      ProcessValue <- "Sequence Times_DB_Dwell Timer_Hours Left"
   IOField "I/O field_66" at 316,321 size 33x28; Authorization "User administration"; FormatPattern 99; Unit d
      ProcessValue <- "Sequence Times_DB_Dwell Timer_Days Left"
   IOField "I/O field_2" at 216,355 size 79x28; Authorization "Commissioning"; FormatPattern 999.9; Unit  Hrs
      ProcessValue <- "Sequence Times_DB_Re-Ox Time"
   IOField "I/O field_67" at 380,355 size 35x28; Authorization "User administration"; FormatPattern 99; Unit m
      ProcessValue <- "Sequence Times_DB_Re-Ox Timer_Minutes Left"
   IOField "I/O field_68" at 348,355 size 33x28; Authorization "User administration"; FormatPattern 99; Unit h
      ProcessValue <- "Sequence Times_DB_Re-Ox Timer_Hours Left"
   IOField "I/O field_69" at 316,355 size 33x28; Authorization "User administration"; FormatPattern 99; Unit d
      ProcessValue <- "Sequence Times_DB_Re-Ox Timer_Days Left"
   IOField "I/O field_70" at 216,389 size 79x28; Authorization "Commissioning"; FormatPattern 999.9; Unit  Hrs
      ProcessValue <- "Sequence Times_DB_Post-Dwell Time"
   IOField "I/O field_71" at 380,389 size 35x28; Authorization "User administration"; FormatPattern 99; Unit m
      ProcessValue <- "Sequence Times_DB_Post-Dwell Timer_Minutes Left"
   IOField "I/O field_72" at 348,389 size 33x28; Authorization "User administration"; FormatPattern 99; Unit h
      ProcessValue <- "Sequence Times_DB_Post-Dwell Timer_Hours Left"
   IOField "I/O field_73" at 316,389 size 33x28; Authorization "User administration"; FormatPattern 99; Unit d
      ProcessValue <- "Sequence Times_DB_Post-Dwell Timer_Days Left"
   Button "Button_1" at 364,1 size 56x38; TextOff 'Text'; PictureOff "Graphic_286"
      on Click: function_efd93a16("Tank Times", 300, 200, -1, -1, 1)
   Group "Group_1" at 20,501 size 235x37

PopupScreen "TANK Activ Warning" 665x250
   Button "Button_1" at 0,0 size 665x250; TextOff 'No TANK Selected. Select a TANK for Tank Treatment.'
      on Release: function_efd93a16("TANK Activ Warning", 300, 200, -1, -1, 1)
   Button "Button_2" at 208,187 size 250x35; TextOff 'OK, Select TANK'
      on Release: ActivateScreen("Balast Water Treatment Setup", 0); function_efd93a16("TANK Activ Warning", 0, 0, -1, -1, 1)

screen "Balast Water Treatment Plant Tank Pressure" 1280x800, template "Template"
   on GenerateScreen: "User_Change"(); "TitleUpdater"()
   Button "HmiScreenItemData_1" at 1,1 size 150x40; TextOn 'Back'; TextOff 'Main Index'
      on Release: ActivateScreen("02 Main Index", 0)
   TextField "Text field_63" at 383,107 size 72x30; Text 'Pre Dwell Time'
   Circle "Circle_29" at 1047,85 size 20x20
      Appearance <- "2102_TIME_CALCS_DB_POST_DWELL_TMR_DN"
   Button "HmiScreenItemData_9" at 10,60 size 158x27; TextOn 'Back'; TextOff 'BWTS Control'
   Button "HmiScreenItemData_4" at 14,150 size 75x47; TextOn 'Back'; TextOff 'Stop'; Authorization "Operate"
      on Release: function_efd93a16("BWTS Stop Confirm", 400, 200, -1, -1, 1)
      ObjectEnable <- "82_To_HMI_CRNT_MODE_GCU"
   Circle "Circle_20" at 137,105 size 29x29
      Appearance <- "80_From_HMI_RUN_IGG(1)"
   Button "HmiScreenItemData_3" at 14,93 size 75x47; TextOn 'Back'; TextOff 'Start'; Authorization "Operate"
      on Release: function_efd93a16("BWTS Start Confirm", 400, 200, -1, -1, 1)
      ObjectEnable <- "82_To_HMI_CRNT_MODE_GCU"
   Button "HmiScreenItemData_2" at 1129,1 size 150x40; TextOn 'Back'; TextOff 'BWTS Setup'
      on Release: ActivateScreen("Balast Water Treatment Setup", 0)
   TextField "Text field_1" at 290,107 size 68x30; Text 'Tank Selected'
   TextField "Text field_2" at 841,107 size 61x30; Text 'BWTS Started'
   TextField "Text field_3" at 568,107 size 62x30; Text 'IGGS Started'
   TextField "Text field_4" at 659,107 size 60x30; Text 'GCU Started'
   TextField "Text field_5" at 748,107 size 61x30; Text 'PGC Started'
   TextField "Text field_6" at 908,107 size 102x30; Text 'Gas Transfer Started'
   Circle "Circle_10" at 956,89 size 14x14
      Appearance <- "2110_BTCS_CNTRL_DB_BTCS_STEP"
   TextField "Text field_7" at 995,107 size 125x30; Text 'Treatment Cycle Completed'
   TextField "Text field_23" at 261,291 size 34x14; Text 'MBG'
   GraphicView "Graphic view_17" at 575,446 size 532x12; Picture "Graphic_151"
   Button "Button_13" at 252,437 size 37x30; TextOff 'DB&B'
   TextField "Text field_58" at 188,226 size 50x40; Text 'Safe Area'
   Button "Button_20" at 724,152 size 115x34; TextOff 'Re-Oxygenation'
      Appearance <- "2110_BTCS_CNTRL_DB_BTCS_STEP"
   Button "Button_21" at 845,152 size 93x34; TextOff 'Post Dwell'
      Appearance <- "2110_BTCS_CNTRL_DB_BTCS_STATE"
   Circle "Circle_1" at 137,105 size 29x29
      Appearance <- "2110_BTCS_CNTRL_DB_BTCS_STATE"
   Circle "Circle_8" at 775,89 size 14x14
      Appearance <- "2110_BTCS_CNTRL_DB_BTCS_STEP"
   Circle "Circle_9" at 685,89 size 14x14
      Appearance <- "100_GCU_AUTO_SEQ_DB_CRNT_STEP"
   Circle "Circle_11" at 595,89 size 14x14
      Appearance <- "51_SLAVE_STATUS_RUNNING"
   Circle "Circle_12" at 866,89 size 14x14
      Appearance <- "2110_BTCS_CNTRL_DB_BTCS_STEP"
   Circle "Circle_13" at 324,89 size 14x14
      Appearance <- "HMI Indication Logic_DB_Tank Selected"
   Circle "Circle_14" at 414,89 size 14x14
      Appearance <- "2102_TIME_CALCS_DB_PRE_DWELL_TMR_DN"
   Button "Button_3" at 626,152 size 93x34; TextOff 'Dwell'
      Appearance <- "2110_BTCS_CNTRL_DB_BTCS_STATE"
   Button "Button_5" at 944,152 size 93x34; TextOff 'Complete'
      Appearance <- "HMI Indication Logic_DB_Sequence Finished"
   TextField "Text field_61" at 202,107 size 71x30; Text 'FA Mode Selected'
   Circle "Circle_2" at 230,89 size 14x14
      Appearance <- "HMI Indication Logic_DB_FA Mode Selected"
   TextField "Text field_60" at 190,519 size 46x25; Text 'GCU'
   GraphicIOField "Graphic I/O field_4" at 187,543 size 53x55; PictureList "GCU"
      ProcessValue <- "100_GCU_AUTO_SEQ_DB_RNG"
   TextField "Text field_74" at 186,279 size 54x25; Text 'IGGS'
   GraphicIOField "Graphic I/O field_1" at 185,303 size 57x53; PictureList "IGGS"
      ProcessValue <- "14_DQ_Data_24PF1"
   TextField "Text field_62" at 183,359 size 60x20; Text 'Disabled'
   TextField "Text field_77" at 183,359 size 60x20; Text 'Enabled'
      Visibility <- "51_SLAVE_STATUS_RUNNING"
   Button "Button_8" at 178,280 size 70x105; TextOff 'Text'
      on Release: ActivateScreen("Inert Gas Generator Plant", 0)
   TextField "Text field_70" at 183,599 size 60x20; Text 'Disabled'
   TextField "Text field_71" at 183,599 size 60x20; Text 'Enabled'
      Visibility <- "100_GCU_AUTO_SEQ_DB_RNG"
   Button "Button_4" at 178,521 size 70x105; TextOff 'Text'
      on Release: ActivateScreen("Inert Gas Conditioning Plant", 0)
   GraphicIOField "Graphic I/O field_2" at 770,45 size 250x30; PictureList "Process time Banner"
      ProcessValue <- "2110_BTCS_CNTRL_DB_BTCS_STATE"
      Visibility <- "2110_BTCS_CNTRL_DB_BTCS_STATE"
   Button "Button_14" at 303,152 size 93x34; TextOff 'Unselected'
      Visibility <- "HMI Indication Logic_DB_Tank Selected"
      Appearance <- "HMI Indication Logic_DB_Tank Selected"
   Button "Button_15" at 404,152 size 93x34; TextOff 'Selected'
      Appearance <- "HMI Indication Logic_DB_Tank Selected"
   Button "Button_16" at 506,152 size 115x34; TextOff 'De-Oxygenation'
      Appearance <- "2110_BTCS_CNTRL_DB_BTCS_STEP"
   TextField "Text field_92" at 304,351 size 76x15; Text 'FIT-418-6P'
   TextField "Text field_98" at 304,308 size 76x15; Text 'FIT-420-6P'
   Button "HmiScreenItemData_19" at 1185,676 size 72x27; TextOn 'Back'; TextOff 'Status'
      on Press: function_efd93a16("Treatment Status", 100, 471, -1, 3, 1)
   Group "Group_6" at 298,44 size 241x30
   Circle "Circle_26" at 504,89 size 14x14
      Appearance <- "2102_TIME_CALCS_DB_Time_To_Treatment"
   TextField "Text field_134" at 470,107 size 75x30; Text 'Wait for IGGS Start'
   GraphicView "Graphic view_4" at 357,210 size 25x62; Picture "Graphic_183"
   GraphicView "Graphic view_5" at 265,210 size 25x62; Picture "Graphic_183"
   IOField "I/O field_31" at 1053,45 size 225x30; FormatPattern ???????????????
      ProcessValue <- "Current User"
   Button "HmiScreenItemData_8" at 772,732 size 503x40; TextOn 'Back'; TextOff 'Text'
   TextField "Screen title" at 783,728 size 496x50; Text 'Screen title'
   Bar "Bar_1" at 262,206 size 122x241; MinimumValue 0; MaximumValue 100
      ProcessValue <- "20_TANKS_IP_DATA_RIO_06_FIRST_TANK_TANKS_PRESS"
   Button "Button_48" at 273,396 size 100x25; TextOff 'DISABLED'
      on Release: function_efd93a16("Tank 6P Status", 168, 315, -1, 2, 1)
      Visibility <- "504_Tank Grouping_DB2020_GROUP of TANK 12"
   Circle "Circle_3" at 340,212 size 14x14
      Appearance <- "20_TANKS_IP_DATA_RIO_06_FIRST_TANK_BWT_LEVEL_HIHI"
   TextField "Text field_125" at 295,212 size 51x14; Text 'LS425-6P'
   Polyline "Polyline_1" at 261,205 size 123x240
      Visibility <- "504_Tank Grouping_DB2020_RUN TANK 12"
   TextField "Text field_64" at 288,273 size 74x20; Text 'Tank - 6P'
   Bar "Bar_2" at 394,206 size 122x241; MinimumValue 0; MaximumValue 100
      ProcessValue <- "20_TANKS_IP_DATA_RIO_05_FIRST_TANK_TANKS_PRESS"
   Button "Button_44" at 406,396 size 100x25; TextOff 'DISABLED'
      on Release: function_efd93a16("Tank 5P Status", 168, 315, -1, 2, 1)
      Visibility <- "504_Tank Grouping_DB2020_GROUP of TANK 10"
   Circle "Circle_4" at 472,212 size 14x14
      Appearance <- "20_TANKS_IP_DATA_RIO_05_FIRST_TANK_BWT_LEVEL_HIHI"
   TextField "Text field_124" at 427,212 size 51x14; Text 'LS425-5P'
   Polyline "Polyline_2" at 392,205 size 123x240
      Visibility <- "504_Tank Grouping_DB2020_RUN TANK 10"
   TextField "Text field_8" at 418,275 size 74x20; Text 'Tank - 5P'
   Bar "Bar_3" at 525,206 size 122x241; MinimumValue 0; MaximumValue 100
      ProcessValue <- "20_TANKS_IP_DATA_RIO_04_FIRST_TANK_TANKS_PRESS"
   Button "Button_40" at 537,395 size 100x25; TextOff 'DISABLED'
      on Release: function_efd93a16("Tank 4P Status", 168, 315, -1, 2, 1)
      Visibility <- "504_Tank Grouping_DB2020_GROUP of TANK 8"
   Circle "Circle_5" at 604,212 size 14x14
      Appearance <- "20_TANKS_IP_DATA_RIO_04_FIRST_TANK_BWT_LEVEL_HIHI"
   TextField "Text field_123" at 559,212 size 51x14; Text 'LS425-4P'
   Polyline "Polyline_3" at 525,205 size 123x240
      Visibility <- "504_Tank Grouping_DB2020_RUN TANK 8"
   TextField "Text field_9" at 553,275 size 74x20; Text 'Tank - 4P'
   Bar "Bar_4" at 657,206 size 122x241; MinimumValue 0; MaximumValue 100
      ProcessValue <- "20_TANKS_IP_DATA_RIO_03_FIRST_TANK_TANKS_PRESS"
   Button "Button_36" at 668,395 size 100x25; TextOff 'DISABLED'
      on Release: function_efd93a16("Tank 3P Status", 168, 315, -1, 0, 1)
      Visibility <- "504_Tank Grouping_DB2020_GROUP of TANK 6"
   Circle "Circle_7" at 736,212 size 14x14
      Appearance <- "20_TANKS_IP_DATA_RIO_03_FIRST_TANK_BWT_LEVEL_HIHI"
   TextField "Text field_122" at 691,212 size 51x14; Text 'LS425-3P'
   Polyline "Polyline_4" at 656,205 size 123x240
      Visibility <- "504_Tank Grouping_DB2020_RUN TANK 6"
   TextField "Text field_14" at 680,275 size 74x20; Text 'Tank - 3P'
   Bar "Bar_5" at 789,206 size 122x241; MinimumValue 0; MaximumValue 100
      ProcessValue <- "20_TANKS_IP_DATA_RIO_02_FIRST_TANK_TANKS_PRESS"
   Button "Button_32" at 802,396 size 100x25; TextOff 'DISABLED'
      on Release: function_efd93a16("Tank 2P Status", 168, 315, -1, 0, 1)
      Visibility <- "504_Tank Grouping_DB2020_GROUP of TANK 4"
   Circle "Circle_15" at 868,212 size 14x14
      Appearance <- "20_TANKS_IP_DATA_RIO_02_FIRST_TANK_BWT_LEVEL_HIHI"
   TextField "Text field_121" at 823,212 size 51x14; Text 'LS425-2P'
   Polyline "Polyline_5" at 789,205 size 123x240
      Visibility <- "504_Tank Grouping_DB2020_RUN TANK 4"
   TextField "Text field_15" at 816,275 size 74x20; Text 'Tank - 2P'
   Bar "Bar_6" at 922,205 size 122x241; MinimumValue 0; MaximumValue 100
      ProcessValue <- "20_TANKS_IP_DATA_RIO_01_FIRST_TANK_TANKS_PRESS"
   Button "Button_52" at 934,395 size 100x25; TextOff 'DISABLED'
      on Release: function_efd93a16("Tank 1P Status", 168, 315, -1, 0, 1)
      Visibility <- "504_Tank Grouping_DB2020_GROUP of TANK 2"
   Circle "Circle_16" at 999,211 size 14x14
      Appearance <- "20_TANKS_IP_DATA_RIO_01_SECOND_TANK_BWT_LEVEL_HIHI"
   TextField "Text field_120" at 955,211 size 51x14; Text 'LS425-1P'
   Polyline "Polyline_6" at 921,205 size 123x240
      Visibility <- "504_Tank Grouping_DB2020_RUN TANK 2"
   GraphicView "Graphic view_6" at 127,446 size 591x12; Picture "Graphic_151"
   TextField "Text field_16" at 947,275 size 74x20; Text 'Tank - 1P'
   Bar "Bar_7" at 1096,334 size 122x241; MinimumValue 0; MaximumValue 100
      ProcessValue <- "20_TANKS_IP_DATA_RIO_01_FIRST_TANK_TANKS_PRESS"
   Circle "Circle_24" at 1168,339 size 14x14
      Appearance <- "20_TANKS_IP_DATA_RIO_01_FIRST_TANK_BWT_LEVEL_HIHI"
   TextField "Text field_133" at 1139,339 size 35x14; Text 'LS425'
   Polyline "Polyline_14" at 1095,332 size 125x242
      Visibility <- "504_Tank Grouping_DB2020_RUN TANK 1"
   Button "Button_56" at 1110,524 size 100x25; TextOff 'DISABLED'
      on Release: function_efd93a16("Tank FP Status", 168, 315, -1, 0, 1)
      Visibility <- "504_Tank Grouping_DB2020_GROUP of TANK 1"
   TextField "Text field_17" at 1111,400 size 111x20; Text 'Fore PeakTank'
   Bar "Bar_8" at 922,458 size 122x258; MinimumValue 0; MaximumValue 100
      ProcessValue <- "20_TANKS_IP_DATA_RIO_01_FIRST_TANK_TANKS_PRESS"
   Button "Button_54" at 933,661 size 100x25; TextOff 'DISABLED'
      on Release: function_efd93a16("Tank 1S Status", 168, 315, -1, 0, 1)
      Visibility <- "504_Tank Grouping_DB2020_GROUP of TANK 3"
   Circle "Circle_23" at 1000,464 size 14x14
      Appearance <- "20_TANKS_IP_DATA_RIO_01_THIRD_TANK_BWT_LEVEL_HIHI"
   TextField "Text field_126" at 955,465 size 51x14; Text 'LS422-1S'
   Polyline "Polyline_7" at 921,458 size 123x259
      Visibility <- "504_Tank Grouping_DB2020_RUN TANK 3"
   TextField "Text field_10" at 950,618 size 74x20; Text 'Tank - 1S'
   Bar "Bar_9" at 790,459 size 122x258; MinimumValue 0; MaximumValue 100
      ProcessValue <- "20_TANKS_IP_DATA_RIO_02_FIRST_TANK_TANKS_PRESS"
   Button "Button_34" at 801,662 size 100x25; TextOff 'DISABLED'
      on Release: function_efd93a16("Tank 2S Status", 168, 315, -1, 0, 1)
      Visibility <- "504_Tank Grouping_DB2020_GROUP of TANK 5"
   Circle "Circle_22" at 868,465 size 14x14
      Appearance <- "20_TANKS_IP_DATA_RIO_02_SECOND_TANK_BWT_LEVEL_HIHI"
   TextField "Text field_127" at 823,466 size 51x14; Text 'LS422-2S'
   Polyline "Polyline_8" at 789,458 size 123x259
      Visibility <- "504_Tank Grouping_DB2020_RUN TANK 5"
   TextField "Text field_11" at 817,618 size 74x20; Text 'Tank - 2S'
   Bar "Bar_10" at 659,460 size 122x258; MinimumValue 0; MaximumValue 100
      ProcessValue <- "20_TANKS_IP_DATA_RIO_03_FIRST_TANK_TANKS_PRESS"
   Button "Button_38" at 669,663 size 100x25; TextOff 'DISABLED'
      on Release: function_efd93a16("Tank 3S Status", 168, 315, -1, 0, 1)
      Visibility <- "504_Tank Grouping_DB2020_GROUP of TANK 7"
   Circle "Circle_21" at 736,467 size 14x14
      Appearance <- "20_TANKS_IP_DATA_RIO_03_SECOND_TANK_BWT_LEVEL_HIHI"
   TextField "Text field_128" at 691,468 size 51x14; Text 'LS422-3S'
   Polyline "Polyline_9" at 658,458 size 123x259
      Visibility <- "504_Tank Grouping_DB2020_RUN TANK 7"
   TextField "Text field_12" at 690,618 size 74x20; Text 'Tank - 3S'
   Bar "Bar_11" at 526,459 size 122x258; MinimumValue 0; MaximumValue 100
      ProcessValue <- "20_TANKS_IP_DATA_RIO_04_FIRST_TANK_TANKS_PRESS"
   Button "Button_42" at 537,662 size 100x25; TextOff 'DISABLED'
      on Release: function_efd93a16("Tank 4S Status", 168, 315, -1, 2, 1)
      Visibility <- "504_Tank Grouping_DB2020_GROUP of TANK 9"
   Circle "Circle_19" at 604,466 size 14x14
      Appearance <- "20_TANKS_IP_DATA_RIO_04_SECOND_TANK_BWT_LEVEL_HIHI"
   TextField "Text field_129" at 559,467 size 51x14; Text 'LS422-4S'
   Polyline "Polyline_10" at 525,458 size 123x259
      Visibility <- "504_Tank Grouping_DB2020_RUN TANK 9"
   TextField "Text field_13" at 554,618 size 74x20; Text 'Tank - 4S'
   Bar "Bar_12" at 394,459 size 122x258; MinimumValue 0; MaximumValue 100
      ProcessValue <- "20_TANKS_IP_DATA_RIO_05_FIRST_TANK_TANKS_PRESS"
   Button "Button_46" at 405,662 size 100x25; TextOff 'DISABLED'
      on Release: function_efd93a16("Tank 5S Status", 168, 315, -1, 2, 1)
      Visibility <- "504_Tank Grouping_DB2020_GROUP of TANK 11"
   Circle "Circle_18" at 472,465 size 14x14
      Appearance <- "20_TANKS_IP_DATA_RIO_05_SECOND_TANK_BWT_LEVEL_HIHI"
   TextField "Text field_130" at 427,466 size 51x14; Text 'LS422-5S'
   Polyline "Polyline_11" at 393,458 size 123x259
      Visibility <- "504_Tank Grouping_DB2020_RUN TANK 11"
   TextField "Text field_18" at 424,618 size 74x20; Text 'Tank - 5S'
   Bar "Bar_13" at 262,460 size 122x258; MinimumValue 0; MaximumValue 100
      ProcessValue <- "20_TANKS_IP_DATA_RIO_06_FIRST_TANK_TANKS_PRESS"
   Button "Button_50" at 273,663 size 100x25; TextOff 'DISABLED'
      on Release: function_efd93a16("Tank 6S Status", 168, 315, -1, 2, 1)
      Visibility <- "504_Tank Grouping_DB2020_GROUP of TANK 13"
   Circle "Circle_17" at 340,467 size 14x14
      Appearance <- "20_TANKS_IP_DATA_RIO_06_SECOND_TANK_BWT_LEVEL_HIHI"
   TextField "Text field_131" at 295,468 size 51x14; Text 'LS422-6S'
   Polyline "Polyline_12" at 261,458 size 123x258
      Visibility <- "504_Tank Grouping_DB2020_RUN TANK 13"
   TextField "Text field_19" at 290,618 size 74x20; Text 'Tank - 6S'
   Bar "Bar_14" at 39,324 size 119x258; Unit %; MinimumValue 0; MaximumValue 100
      ProcessValue <- "20_TANKS_IP_DATA_RIO_07_FIRST_TANK_TANKS_PRESS"
   Circle "Circle_25" at 108,330 size 14x14
      Appearance <- "20_TANKS_IP_DATA_RIO_07_FIRST_TANK_BWT_LEVEL_HIHI"
   TextField "Text field_132" at 79,330 size 35x14; Text 'LS425'
   Polyline "Polyline_13" at 38,324 size 121x259
      Visibility <- "504_Tank Grouping_DB2020_RUN TANK 14"
   Button "Button_58" at 48,527 size 100x25; TextOff 'DISABLED'
      on Release: function_efd93a16("Tank AP Status", 168, 315, -1, 2, 1)
      Visibility <- "504_Tank Grouping_DB2020_GROUP of TANK 14"
   Button "HmiScreenItemData_6" at 1043,144 size 116x50; TextOn 'Back'; TextOff 'Tank Status'
      on Release: ActivateScreen("Balast Water Treatment Plant", 0)
   Button "Button_2" at 252,437 size 37x30; TextOff 'DB&B'
      on Release: function_efd93a16("Double Block & Bleed Valve Monitoring", 250, 250, -1, -1, 1)
      Appearance <- "10_DI_DATA_CV407_OPN"
   TextField "Text field_65" at 190,398 size 46x25; Text 'PGC'
   TextField "Text field_75" at 183,480 size 60x20; Text 'Disabled'
   TextField "Text field_76" at 183,480 size 60x20; Text 'Enabled'
      Visibility <- "10_DI_DATA_E_400_RUN"
   GraphicView "Graphic view_76" at 185,421 size 57x55; Picture "Graphic_251"
   Button "Button_6" at 179,402 size 70x105; TextOff 'Text'
      on Release: ActivateScreen("PGC System", 0)
   TextField "Text field_20" at 53,396 size 103x20; Text 'Aft PeakTank'
   GraphicView "Graphic view_108" at 4,683 size 96x48; Picture "Left Arow"
   Button "HmiScreenItemData_14" at 3,660 size 106x93; TextOn 'Back'; TextOff 'Text'
      on Press: ActivateScreen("Inert Gas Conditioning Plant", 0)
   IOField "I/O field_1" at 44,460 size 115x25; FormatPattern s999.9; Unit mBar
      ProcessValue <- "20_TANKS_IP_DATA_RIO_07_FIRST_TANK_TANKS_PRESS"
   IOField "I/O field_2" at 269,331 size 114x25; FormatPattern s999.9; Unit mBar
      ProcessValue <- "20_TANKS_IP_DATA_RIO_06_FIRST_TANK_TANKS_PRESS"
   IOField "I/O field_3" at 398,331 size 117x25; FormatPattern s999.9; Unit mBar
      ProcessValue <- "20_TANKS_IP_DATA_RIO_05_FIRST_TANK_TANKS_PRESS"
   IOField "I/O field_4" at 531,331 size 117x25; FormatPattern s999.9; Unit mBar
      ProcessValue <- "20_TANKS_IP_DATA_RIO_04_FIRST_TANK_TANKS_PRESS"
   IOField "I/O field_5" at 662,331 size 114x25; FormatPattern s999.9; Unit mBar
      ProcessValue <- "20_TANKS_IP_DATA_RIO_03_FIRST_TANK_TANKS_PRESS"
   IOField "I/O field_6" at 796,331 size 119x25; FormatPattern s999.9; Unit mBar
      ProcessValue <- "20_TANKS_IP_DATA_RIO_02_FIRST_TANK_TANKS_PRESS"
   IOField "I/O field_7" at 928,331 size 118x25; FormatPattern s999.9; Unit mBar
      ProcessValue <- "20_TANKS_IP_DATA_RIO_01_FIRST_TANK_TANKS_PRESS"
   IOField "I/O field_8" at 1103,459 size 119x25; FormatPattern s999.9; Unit mBar
      ProcessValue <- "20_TANKS_IP_DATA_RIO_01_FIRST_TANK_TANKS_PRESS"
   IOField "I/O field_9" at 928,555 size 118x25; FormatPattern s999.9; Unit mBar
      ProcessValue <- "20_TANKS_IP_DATA_RIO_01_FIRST_TANK_TANKS_PRESS"
   IOField "I/O field_10" at 796,556 size 118x25; FormatPattern s999.9; Unit mBar
      ProcessValue <- "20_TANKS_IP_DATA_RIO_02_FIRST_TANK_TANKS_PRESS"
   IOField "I/O field_11" at 664,558 size 116x25; FormatPattern s999.9; Unit mBar
      ProcessValue <- "20_TANKS_IP_DATA_RIO_03_FIRST_TANK_TANKS_PRESS"
   IOField "I/O field_12" at 530,557 size 117x25; FormatPattern s999.9; Unit mBar
      ProcessValue <- "20_TANKS_IP_DATA_RIO_04_FIRST_TANK_TANKS_PRESS"
   IOField "I/O field_13" at 400,558 size 114x25; FormatPattern s999.9; Unit mBar
      ProcessValue <- "20_TANKS_IP_DATA_RIO_05_FIRST_TANK_TANKS_PRESS"
   IOField "I/O field_14" at 268,559 size 116x25; FormatPattern s999.9; Unit mBar
      ProcessValue <- "20_TANKS_IP_DATA_RIO_06_FIRST_TANK_TANKS_PRESS"
   Button "Button_88" at 34,324 size 127x264; TextOff 'Text'
      on Release: function_efd93a16("Tank AP Status", 168, 315, -1, 0, 1)
      Appearance <- "504_Tank Grouping_DB2020_RUN TANK 14"
   Button "Button_86" at 259,458 size 126x260; TextOff 'Text'
      on Release: function_efd93a16("Tank 6S Status", 168, 315, -1, 0, 1)
      Appearance <- "504_Tank Grouping_DB2020_RUN TANK 13"
   Button "Button_79" at 391,457 size 126x262; TextOff 'Text'
      on Release: function_efd93a16("Tank 5S Status", 168, 315, -1, 0, 1)
      Appearance <- "504_Tank Grouping_DB2020_RUN TANK 11"
   Button "Button_77" at 523,457 size 126x262; TextOff 'Text'
      on Release: function_efd93a16("Tank 4S Status", 168, 315, -1, 0, 1)
      Appearance <- "504_Tank Grouping_DB2020_RUN TANK 9"
   Button "Button_74" at 657,457 size 126x262; TextOff 'Text'
      on Release: function_efd93a16("Tank 3S Status", 168, 315, -1, 0, 1)
      Appearance <- "504_Tank Grouping_DB2020_RUN TANK 7"
   Button "Button_70" at 788,457 size 126x262; TextOff 'Text'
      on Release: function_efd93a16("Tank 2S Status", 168, 315, -1, 0, 1)
      Appearance <- "504_Tank Grouping_DB2020_RUN TANK 5"
   Button "Button_66" at 921,457 size 126x261; TextOff 'Text'
      on Release: function_efd93a16("Tank 1S Status", 168, 315, -1, 0, 1)
      Appearance <- "504_Tank Grouping_DB2020_RUN TANK 3"
   Button "Button_61" at 1093,328 size 130x248; TextOff 'Text'
      on Release: function_efd93a16("Tank FP Status", 168, 315, -1, 0, 1)
      Appearance <- "504_Tank Grouping_DB2020_RUN TANK 1"
   Button "Button_62" at 919,205 size 126x242; TextOff 'Text'
      on Release: function_efd93a16("Tank 1P Status", 168, 315, -1, 0, 1)
      Appearance <- "504_Tank Grouping_DB2020_RUN TANK 2"
   Button "Button_68" at 789,202 size 126x246; TextOff 'Text'
      on Release: function_efd93a16("Tank 2P Status", 168, 315, -1, 0, 1)
      Appearance <- "504_Tank Grouping_DB2020_RUN TANK 4"
   Button "Button_72" at 654,205 size 126x242; TextOff 'Text'
      on Release: function_efd93a16("Tank 3P Status", 168, 315, -1, 0, 1)
      Appearance <- "504_Tank Grouping_DB2020_RUN TANK 6"
   Button "Button_76" at 524,205 size 126x243; TextOff 'Text'
      on Release: function_efd93a16("Tank 4P Status", 168, 315, -1, 0, 1)
      Appearance <- "504_Tank Grouping_DB2020_RUN TANK 8"
   Button "Button_78" at 392,206 size 126x241; TextOff 'Text'
      on Release: function_efd93a16("Tank 5P Status", 168, 315, -1, 0, 1)
      Appearance <- "504_Tank Grouping_DB2020_RUN TANK 10"
   Button "Button_84" at 259,204 size 126x244; TextOff 'Text'
      on Release: function_efd93a16("Tank 6P Status", 168, 315, -1, 0, 1)
      Appearance <- "504_Tank Grouping_DB2020_RUN TANK 12"
   Group "Group_5" at 664,46 size 45x27; FormatPattern 999
   Group "Group_1" at 711,46 size 50x27; FormatPattern 999; Unit h
   Group "Group_2" at 605,46 size 57x27; FormatPattern 999; Unit h
   Button "HmiScreenItemData_5" at 180,144 size 116x50; TextOn 'Back'; TextOff 'Tank Status'
      on Release: function_efd93a16("Tank Status", 400, 250, -1, -1, 1)
   Button "Button_10" at 14,93 size 153x55; TextOff 'Text'
      on Release: function_efd93a16("Salinity - Acceptance", 168, 315, -1, 0, 1)
      Visibility <- "2068_Sys_Status_Data_SAL_VALID"
   Button "Button_12" at 14,93 size 153x53; TextOff 'Text'
      on Release: function_efd93a16("Tank Times", 300, 200, -1, 0, 1)
      Visibility <- "2068_Sys_Status_Data_Times Visibil"
   Button "Button_59" at 298,44 size 240x30; TextOn 'TB3 Enabled'; TextOff 'BWT System Shutting Down'
      Visibility <- "2110_BTCS_CNTRL_DB_BTCS_STATE"
   Button "Button_60" at 299,44 size 240x30; TextOn 'TB3 Enabled'; TextOff 'BWT System Enabled'
      Visibility <- "2110_BTCS_CNTRL_DB_BTCS_STATE"
   IOField "I/O field_29" at 664,46 size 45x27; FormatPattern 99; Unit h
      Visibility <- "2110_BTCS_CNTRL_DB_BTCS_STATE"
      ProcessValue <- "Sequence Times_DB_Treatment Timer_Hours Left"
   IOField "I/O field_30" at 664,46 size 45x27; FormatPattern 99; Unit h
      Visibility <- "2110_BTCS_CNTRL_DB_BTCS_STATE"
      ProcessValue <- "Sequence Times_DB_Pre-Dwell Timer_Hours Left"
   IOField "I/O field_15" at 711,46 size 50x27; FormatPattern 99; Unit m
      Visibility <- "2110_BTCS_CNTRL_DB_BTCS_STATE"
      ProcessValue <- "Sequence Times_DB_Treatment Timer_Minutes Left"
   IOField "I/O field_16" at 711,46 size 50x27; FormatPattern 99; Unit m
      Visibility <- "2110_BTCS_CNTRL_DB_BTCS_STATE"
      ProcessValue <- "Sequence Times_DB_Pre-Dwell Timer_Minutes Left"
   IOField "I/O field_17" at 605,46 size 57x27; FormatPattern 999; Unit d
      Visibility <- "2110_BTCS_CNTRL_DB_BTCS_STATE"
      ProcessValue <- "Sequence Times_DB_Treatment Timer_Days Left"
   IOField "I/O field_18" at 605,46 size 57x27; FormatPattern 999; Unit d
      Visibility <- "2110_BTCS_CNTRL_DB_BTCS_STATE"
      ProcessValue <- "Sequence Times_DB_Pre-Dwell Timer_Days Left"

VB script "BWT_Warning"
   If SmartTags("2068_Sys_Status_Data_Not BWT mode Warning") Then
   	efd93a16-2665-4b85-bcb9-25eddcb7b6f4 BWT Mode Warning,275,250,$3$hmiOn$,$3$hmiTop$,$3$hmiMedium$
   'ElseIf Not SmartTags("BWT Mode Warning") Then
   '	ShowPopupScreen"BWT Mode Warning",0,0,hmiOff,hmiAnimationOff,hmiMedium
   End If

VB script "PGCCommissioning"
   If SmartTags("PGC_COMMISSION_MODE_DB_Drive Popup") Then
   	efd93a16-2665-4b85-bcb9-25eddcb7b6f4 PGC Commissioning, 0, 0, $3$hmiOn$, $3$hmiBottom$, $3$hmiMedium$
   	ElseIf Not SmartTags("PGC_COMMISSION_MODE_DB_Drive Popup") Then
   efd93a16-2665-4b85-bcb9-25eddcb7b6f4 PGC Commissioning, 0, 0, $3$hmiOff$, $3$hmiOff$, $3$hmiMedium$
   End If

VB script "HeartBeatFunction"
   If SmartTags("CCR HMI HEART BEAT")=0 Then
   	b21d3eaf-4e31-425c-ad1a-ba4e4002cacc(CCR HMI HEART BEAT),1
   Else
   	b21d3eaf-4e31-425c-ad1a-ba4e4002cacc (CCR HMI HEART BEAT),0
   End If

VB script "Salinity_FreshWaterAlert"
   If SmartTags("2068_Sys_Status_Data_SAL_CNF_CHK") Then
   	efd93a16-2665-4b85-bcb9-25eddcb7b6f4 Salinity - Fresh Water Alert,789,316,$3$hmiOn$,$3$hmiBottom$,$3$hmiMedium$
   ElseIf Not SmartTags("2068_Sys_Status_Data_SAL_CNF_CHK") Then
   	efd93a16-2665-4b85-bcb9-25eddcb7b6f4Salinity - Fresh Water Alert,0,0,$3$hmiOff$,$3$hmiAnimationOff$,$3$hmiMedium$
   End If

VB script "SD_Card_Overflow"
   If SmartTags("Logging SD Card Overflow") Then 
   	efd93a16-2665-4b85-bcb9-25eddcb7b6f4 SD Card overflow,275,250,$3$hmiOn$,$3$hmiBottom$,$3$hmiMedium$
   ElseIf Not SmartTags("Logging SD Card Overflow") Then
   	efd93a16-2665-4b85-bcb9-25eddcb7b6f4SD Card overflow,0,0,$3$hmiOff$,$3$hmiAnimationOff$,$3$hmiMedium$
   End If

VB script "TimeRemainingToTreatment"
   If SmartTags("Warn To Start IGG") Then
   	efd93a16-2665-4b85-bcb9-25eddcb7b6f4 Time Until Treatment Required, 400, 200, $3$hmiOn$, $3$hmiBottom$, $3$hmiMedium$
   	ElseIf Not SmartTags("Warn To Start IGG") Then
   efd93a16-2665-4b85-bcb9-25eddcb7b6f4 Time Until Treatment Required, 0, 0, $3$hmiOff$, $3$hmiOff$, $3$hmiMedium$
   End If

VB script "TitleUpdater"
   Dim title
   Set title = HmiRuntime.ActiveScreen.ScreenItems("Screen title")
   title.Text = HmiRuntime.ActiveScreen.ObjectName

VB script "TreatmentCycleCompleted"
   If SmartTags("Sequence Times_DB_Post-Dwell Timer_Q") Then
   	efd93a16-2665-4b85-bcb9-25eddcb7b6f4 Treatment Cycle Completed,275,250,$3$hmiOn$,$3$hmiBottom$,$3$hmiMedium$
   'ElseIf Not SmartTags("Treatment Runs Completed") Then
   '	ShowPopupScreen"Treatment Cycle Completed",0,0,hmiOff,hmiAnimationOff,hmiMedium
   End If

VB script "TreatmentdDailyChecks"
   If SmartTags("88_treatment_POP_UP") Then
   	efd93a16-2665-4b85-bcb9-25eddcb7b6f4 Treatment check / Daily Checks Completed,275,250,$3$hmiOn$,$3$hmiBottom$,$3$hmiMedium$
   End If

VB script "TreatmentRequired"
   If SmartTags("Warn To Start IGG-Last") Then
   	efd93a16-2665-4b85-bcb9-25eddcb7b6f4 Start Treatment, 400, 200, $3$hmiOn$, $3$hmiBottom$, $3$hmiMedium$
   	ElseIf Not SmartTags("Warn To Start IGG-Last") Then
       efd93a16-2665-4b85-bcb9-25eddcb7b6f4 Start Treatment, 0, 0, $3$hmiOff$, $3$hmiOff$, $3$hmiMedium$
   End If

VB script "User_Change"
   f41c6f6c-971d-4734-9362-16d81ac70597 Current User
   e1ab61de-e5a2-437b-97c4-abda991a3a2e user_group
   
   'Tip:
   ' 1. Use the <CTRL+SPACE> or <CTRL+I> shortcut to open a list of all objects and functions
   ' 2. Write the code using the HMI Runtime object.
   '  Example: HmiRuntime.Screens("Screen_1").
   ' 3. Use the <CTRL+J> shortcut to create an object reference.
   'Write the code as of this position:

VB script "VoyageTimeInsufficient"
   If SmartTags("Voyage Time Invalid") Then
   	efd93a16-2665-4b85-bcb9-25eddcb7b6f4 Voyage Time Warning,275,250,$3$hmiOn$,$3$hmiTop$,$3$hmiMedium$
   ElseIf Not SmartTags("Voyage Time Invalid") Then
   	efd93a16-2665-4b85-bcb9-25eddcb7b6f4Voyage Time Warning,0,0,$3$hmiOff$,$3$hmiAnimationOff$,$3$hmiMedium$
   End If

VB script "ALARM_Present"
   If SmartTags("60_Alarm_Data_ALRM_PRSNT") Then
   	bec8f1e5-2ab1-45f6-ad91-1d37c469eb91 04 Alarm Log,0
   End If
   
   'If Not SmartTags("60_Alarm_Data_ALRM_PRSNT") Then
   '	ActivateScreen "01 Home",0
   'End If
   
   
   
   
   
   
   
   
   
   'Tip:
   ' 1. Use the <CTRL+SPACE> or <CTRL+I> shortcut to open a list of all objects and functions
   ' 2. Write the code using the HMI Runtime object.
   '  Example: HmiRuntime.Screens("Screen_1").
   ' 3. Use the <CTRL+J> shortcut to create an object reference.
   'Write the code as of this position:

VB script "HeartBeatHMI_Warning"
   Dim Warning, Tempos
   
   
   If SmartTags("HEART BEAT TRUE")=True Then
   	Warning=0 '"HEART BEAT TRUE"
   Else
   	Warning=1
   End If
   
   If Warning=0 Then
   	efd93a16-2665-4b85-bcb9-25eddcb7b6f4 Lost Comunication, 0, 0, $3$hmiOff$, $3$hmiOff$, $3$hmiMedium$
   Else
   	efd93a16-2665-4b85-bcb9-25eddcb7b6f4 Lost Comunication, 300, 100, $3$hmiOn$, $3$hmiBottom$, $3$hmiMedium$
   End If		
   
   	b21d3eaf-4e31-425c-ad1a-ba4e4002cacc SmartTags("HEART BEAT TRUE"),False

VB script "PGC_ProtectionWarning"
   If SmartTags("Setpoint Override_DB_Set Pressure") Then
   	efd93a16-2665-4b85-bcb9-25eddcb7b6f4 PGC Protection Warning,275,200,$3$hmiOn$,$3$hmiTop$,$3$hmiMedium$
   'ElseIf Not SmartTags("Setpoint Override_DB_Set Pressure") Then
   '	ShowPopupScreen"Setpoint Override_DB_Set Pressure",0,0,hmiOff,hmiAnimationOff,hmiMedium
   End If

VB script "TreatmentRequired_GCU"
   If SmartTags("Warn To Start GCU-Last") Then
   	efd93a16-2665-4b85-bcb9-25eddcb7b6f4 Start GCU for Re-Ox, 400, 200, $3$hmiOn$, $3$hmiBottom$, $3$hmiMedium$
   	ElseIf Not SmartTags("Warn To Start GCU-Last") Then
   efd93a16-2665-4b85-bcb9-25eddcb7b6f4 Start GCU for Re-Ox, 0, 0, $3$hmiOff$, $3$hmiOff$, $3$hmiMedium$
   End If

VB script "TimeRemainingToRe_Ox"
   If SmartTags("Warn To Start GCU") Then
   	efd93a16-2665-4b85-bcb9-25eddcb7b6f4 Time Until GCU Start Required, 400, 200, $3$hmiOn$, $3$hmiBottom$, $3$hmiMedium$
   	ElseIf Not SmartTags("Warn To Start GCU") Then
   efd93a16-2665-4b85-bcb9-25eddcb7b6f4 Time Until GCU Start Required, 0, 0, $3$hmiOff$, $3$hmiOff$, $3$hmiMedium$
   End If

VB script "TANK_Activ_Warning"
   If SmartTags("Not TANK Activ Warning") Then
   	efd93a16-2665-4b85-bcb9-25eddcb7b6f4 TANK Activ Warning,300,200,$3$hmiOn$,$3$hmiTop$,$3$hmiMedium$
   'ElseIf Not SmartTags("Not TANK Activ Warning") Then
   '	ShowPopupScreen"TANK Activ Warning",0,0,hmiOff,hmiAnimationOff,hmiMedium
   End If

scheduled task "VB procces"
   Triggers <- "1 min"

scheduled task "User Change"
   on Action: "User_Change"()

scheduled task "Heart Beat"
   on Action: "HeartBeatFunction"(); "HeartBeatHMI_Warning"()
   Triggers <- "1 min"
*)

(* ===== HMI "HMI_RT_2" =====
system functions are stored by id; their names below are inferred from use
connection "IGG PLC Comms_1": ETHERNET, S7_1500_OMS
connection "BC PLC Comms_1": ETHERNET, S7_1500_OMS
connection "BWTS PLC Comms_1": ETHERNET, S7_1500_OMS

